// TIA Portal project "liquid refill system" (V18)

(* hardware
DEVICE "S7-1200 station_1"  S7-1200 Station
   slot 0: "Rack_0"  S7-1200 Rack  Rack  V1.0
   slot 1: "PLC_Refill"  CPU 1214C DC/DC/Rly  6ES7 214-1HG40-0XB0  V4.6
DEVICE "HMI_Refill"  TP900 Comfort
   slot 0: "HMI_Refill"  TP900 Comfort  6AV2 124-0JC01-0AX0  17.0.0.0
   slot 1: "HMI_RT_1"  TP900 Comfort  6AV2 124-0JC01-0AX0  17.0.0.0
   slot 5: "HMI_Refill.IE_CP_1"  PROFINET Interface  17.0.0.0
      slot 1: "PROFINET Interface_1"  PROFINET Interface
         slot 1: "Port_1"  Port
         slot 2: "Port_2"  Port
   slot 7: "HMI_Refill.MPI/DP_CP_1"  MPI/DP Interface  17.0.0.0
*)

// ===== PLC "PLC_Refill"  CPU 1214C DC/DC/Rly =====

VAR_GLOBAL   // PLC tag table "Default tag table"
   "System_Byte" AT %MB1 : Byte;
   "FirstScan" AT %M1.0 : Bool;
   "DiagStatusUpdate" AT %M1.1 : Bool;
   "AlwaysTRUE" AT %M1.2 : Bool;
   "AlwaysFALSE" AT %M1.3 : Bool;
   "Clock_Byte" AT %MB0 : Byte;
   "Clock_10Hz" AT %M0.0 : Bool;
   "Clock_5Hz" AT %M0.1 : Bool;
   "Clock_2.5Hz" AT %M0.2 : Bool;
   "Clock_2Hz" AT %M0.3 : Bool;
   "Clock_1.25Hz" AT %M0.4 : Bool;
   "Clock_1Hz" AT %M0.5 : Bool;
   "Clock_0.625Hz" AT %M0.6 : Bool;
   "Clock_0.5Hz" AT %M0.7 : Bool;
END_VAR

VAR_GLOBAL   // PLC tag table "input Machine"
   "i_Start" AT %I0.0 : Bool;
   "i_Stop" AT %I0.1 : Bool;
   "i_Reset" AT %I0.2 : Bool;
END_VAR

VAR_GLOBAL   // PLC tag table "output Machine"
   "q_Lamp_Running" AT %Q0.0 : Bool;   // Indication lamp, application running
   "q_Lamp_Faulted" AT %Q0.1 : Bool;   // Indication lamp, application faulted
   "q_Lamp_Ready" AT %Q0.7 : Bool;   // Indication lamp, application ready
END_VAR

VAR_GLOBAL   // PLC tag table "input Equipment"
   "iw_RefillTank1_Level" AT %IW64 : Int;   // Refill tank actual water level process
   "iw_RefillTank2_Level" AT %IW66 : Int;   // Refill tank actual water level process
   "i_RefillPump1_MCB" AT %I0.3 : Bool;   // Refill pump motor circuit breaker process ( Motor saftety )
   "i_RefillPump1_LI" AT %I0.4 : Bool;   // Refill pump local isolator process( Human safety )
   "i_RefillPump1_running" AT %I0.5 : Bool;   // Refill Pump Running feedback
   "i_RefillValve1_feedback" AT %I0.6 : Bool;   // Refill Valve position open feedback
   "i_RefillPump2_MCB" AT %I0.7 : Bool;   // Refill pump motor circuit breaker process ( Motor saftety )
   "i_RefillPump2_LI" AT %I1.0 : Bool;   // Refill pump local isolator process( Human safety )
   "i_RefillPump2_running" AT %I1.1 : Bool;   // Refill Pump Running feedback
   "i_RefillValve2_feedback" AT %I1.2 : Bool;   // Refill Valve position open feedback
   "i_SupplyTank_lowlevel" AT %I1.3 : Bool;   // Supply tank low level indicator
   "i_SupplyValve_feedback" AT %I1.4 : Bool;   // Supply valve position open feedback
END_VAR

VAR_GLOBAL   // PLC tag table "output Equipment"
   "q_RefillPump1_Start" AT %Q0.2 : Bool;   // Refill pump start operation process
   "q_RefillValve1_Open" AT %Q0.3 : Bool;   // Refill valve open operation process
   "q_RefillPump2_Start" AT %Q0.4 : Bool;   // Refill pump start operation process
   "q_RefillValve2_Open" AT %Q0.5 : Bool;   // Refill valve open operation process
   "q_SupplyValve_Open" AT %Q0.6 : Bool;   // Supply valve open operation process
END_VAR

TYPE "UDT_Statehandler"
   STRUCT
      State : Struct   // System states
         iState : Int;   // State feedback
         xReady : Bool;   // System is in ready state
         xRunning : Bool;   // System is in running state
         xFaulted : Bool;   // System is in faulted state
         xReset : Bool;   // System is in reset fault state
      END_STRUCT;
      Cmd : Struct   // Command structure
         xStart : Bool;   // Start operation - button on HMI
         xStop : Bool;   // Stop operation - button on HMI
         xReset : Bool;   // Reset faults - button on HMI
      END_STRUCT;
   END_STRUCT;
END_TYPE

TYPE "UDT_Refill"
   STRUCT
      Sts : Struct   // Status structure
         iTankLevel : Int;   // Actual product level in tank
         iPumpState : Int;   // Pump state (0=off,1=running,2=faulted)
         iValveState : Int;   // Valve state (0=closed,1=open,2=faulted)
         xPumpRunning : Bool;   // Pump is in operation
         xValveOpen : Bool;   // Valve is in open position
         xFaulted : Bool;   // Refill system faulted
      END_STRUCT;
      Cmd : Struct   // Command structure
         xRequestRefill : Bool;   // Request a refill
      END_STRUCT;
      Par : Struct   // Parameter structure
         iTankLevelLow : Int;   // Tank low level (%)
         iTankLevelHigh : Int;   // Tank high level (%)
      END_STRUCT;
      Cfg : Struct   // Configuration structure
         xSpare : Bool;   // spare ( reserve )
      END_STRUCT;
      Flt : Struct   // Fault Structure
         wTrigger : Word;   // Fault triggers
      END_STRUCT;
   END_STRUCT;
END_TYPE

TYPE "UDT_Supply"
   STRUCT
      Sts : Struct   // Status structure
         iValveState : Int;   // Valve state (0=closed,1=open,2=faulted)
         xTankLowLevel : Bool;   // Low product level in tank
         xValveOpen : Bool;   // Valve is in open position
         xFaulted : Bool;   // Supply system faulted
      END_STRUCT;
      Cmd : Struct   // Command structure
         xSpare : Bool;   // spare(reserve)
      END_STRUCT;
      Par : Struct   // Parameter structure
         rTankLowLevelDelay : Real;   // rTankLowLevelDelay
      END_STRUCT;
      Cfg : Struct   // Configuration structure
         xSpare : Bool;   // spare(reserve)
      END_STRUCT;
      Flt : Struct   // Fault structure
         wTrigger : Word;   // Fault triggers
      END_STRUCT;
   END_STRUCT;
END_TYPE

// folder: 00 Machine

DATA_BLOCK "Instance_Machine Module"   // DB4
{ S7_Optimized_Access := 'TRUE' }
VERSION : 0.1
// stored: InstanceOfName FB_Machine Module
"FB_Machine Module"
BEGIN
END_DATA_BLOCK

// folder: 01 Equipment

DATA_BLOCK "FB_Equipment Modules_DB"   // DB5
{ S7_Optimized_Access := 'TRUE' }
VERSION : 0.1
// stored: InstanceOfName FB_Equipment Modules
"FB_Equipment Modules"
BEGIN
END_DATA_BLOCK

// folder: Global DB

DATA_BLOCK "DB - Machine"   // DB1
{ S7_Optimized_Access := 'TRUE' }
VERSION : 0.1
   VAR
      StateHandler : "UDT_Statehandler";
   END_VAR
BEGIN
END_DATA_BLOCK

DATA_BLOCK "DB - Equipment"   // DB2
{ S7_Optimized_Access := 'TRUE' }
VERSION : 0.1
   VAR
      Supply : "UDT_Supply";
      Refill_Process_1 : "UDT_Refill";
      Refill_Process_2 : "UDT_Refill";
   END_VAR
BEGIN
END_DATA_BLOCK

// folder: (top level)

ORGANIZATION_BLOCK "Main"   // OB1, LAD, ProgramCycle
TITLE = "Main Program Sweep (Cycle)"
{ S7_Optimized_Access := 'TRUE' }
VERSION : 0.1
   VAR_INPUT
      Initial_Call : Bool;   // Initial call of this OB
      Remanence : Bool;   // =True, if remanent data are available
   END_VAR
BEGIN

REGION Network 1: CALL - Main machine modules
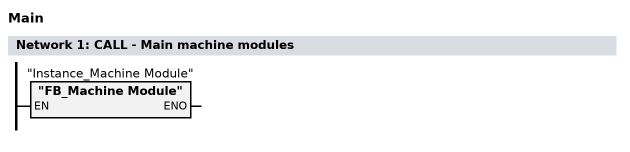
   RUNG wire#powerrail
      "Instance_Machine Module"()
   END_RUNG
   // the same network as SCL:
   "Instance_Machine Module"();   // "FB_Machine Module"
END_REGION

REGION Network 2: CALL - Main equipment modules
END_REGION
END_ORGANIZATION_BLOCK

// folder: 00 Machine

FUNCTION_BLOCK "FB_Machine Module"   // FB1, LAD
{ S7_Optimized_Access := 'TRUE' }
VERSION : 0.1
   VAR
      FB_StateHandler_Instance : "FB_StateHandler";
   END_VAR
   VAR_TEMP
      info : Struct
         xReady : Bool;
         xRunning : Bool;
         xFaulted : Bool;
         xReset : Bool;
      END_STRUCT;
   END_VAR
BEGIN

REGION Network 1
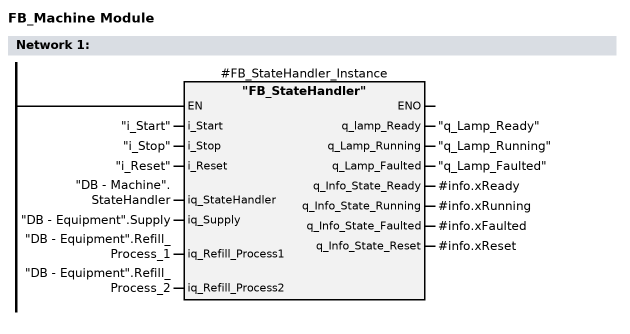
   RUNG wire#powerrail
      #FB_StateHandler_Instance(i_Start := "i_Start", i_Stop := "i_Stop", i_Reset := "i_Reset", iq_StateHandler := "DB - Machine".StateHandler, iq_Supply := "DB - Equipment".Supply, iq_Refill_Process1 := "DB - Equipment".Refill_Process_1, iq_Refill_Process2 := "DB - Equipment".Refill_Process_2, q_lamp_Ready => "q_Lamp_Ready", q_Lamp_Running => "q_Lamp_Running", q_Lamp_Faulted => "q_Lamp_Faulted", q_Info_State_Ready => #info.xReady, q_Info_State_Running => #info.xRunning, q_Info_State_Faulted => #info.xFaulted, q_Info_State_Reset => #info.xReset)
   END_RUNG
   // the same network as SCL:
   #FB_StateHandler_Instance(i_Start := "i_Start",   // "FB_StateHandler"
                           i_Stop := "i_Stop",
                           i_Reset := "i_Reset",
                           iq_StateHandler := "DB - Machine".StateHandler,
                           iq_Supply := "DB - Equipment".Supply,
                           iq_Refill_Process1 := "DB - Equipment".Refill_Process_1,
                           iq_Refill_Process2 := "DB - Equipment".Refill_Process_2,
                           q_lamp_Ready => "q_Lamp_Ready",
                           q_Lamp_Running => "q_Lamp_Running",
                           q_Lamp_Faulted => "q_Lamp_Faulted",
                           q_Info_State_Ready => #info.xReady,
                           q_Info_State_Running => #info.xRunning,
                           q_Info_State_Faulted => #info.xFaulted,
                           q_Info_State_Reset => #info.xReset);
END_REGION
END_FUNCTION_BLOCK

// folder: 00 Machine/Function

FUNCTION_BLOCK "FB_StateHandler"   // FB2, LAD
TITLE = MACHINE - State Handler
{ S7_Optimized_Access := 'TRUE' }
VERSION : 0.1
// This function block contains all logic for control and status of the machine state handler.
// This module consists of 4 states: start, stop, faulted and reset.
   VAR_INPUT
      i_Start : Bool;
      i_Stop : Bool;
      i_Reset : Bool;
   END_VAR
   VAR_OUTPUT
      q_lamp_Ready : Bool;
      q_Lamp_Running : Bool;   // Lamp machine running
      q_Lamp_Faulted : Bool;   // Lamp machine faulted
      q_Info_State_Ready : Bool;
      q_Info_State_Running : Bool;
      q_Info_State_Faulted : Bool;
      q_Info_State_Reset : Bool;
   END_VAR
   VAR_IN_OUT
      iq_StateHandler : "UDT_Statehandler";
      iq_Supply : "UDT_Supply";
      iq_Refill_Process1 : "UDT_Refill";
      iq_Refill_Process2 : "UDT_Refill";
   END_VAR
   VAR
      stOnDelay_Reset : IEC_TIMER;
      iState : Int;
   END_VAR
   VAR_TEMP
      _tTimeET : Time;
   END_VAR
BEGIN

REGION Network 1: CONTROL - Start Operation
   // The application goes from a ready state (0) to a running state (1) by pressing Start
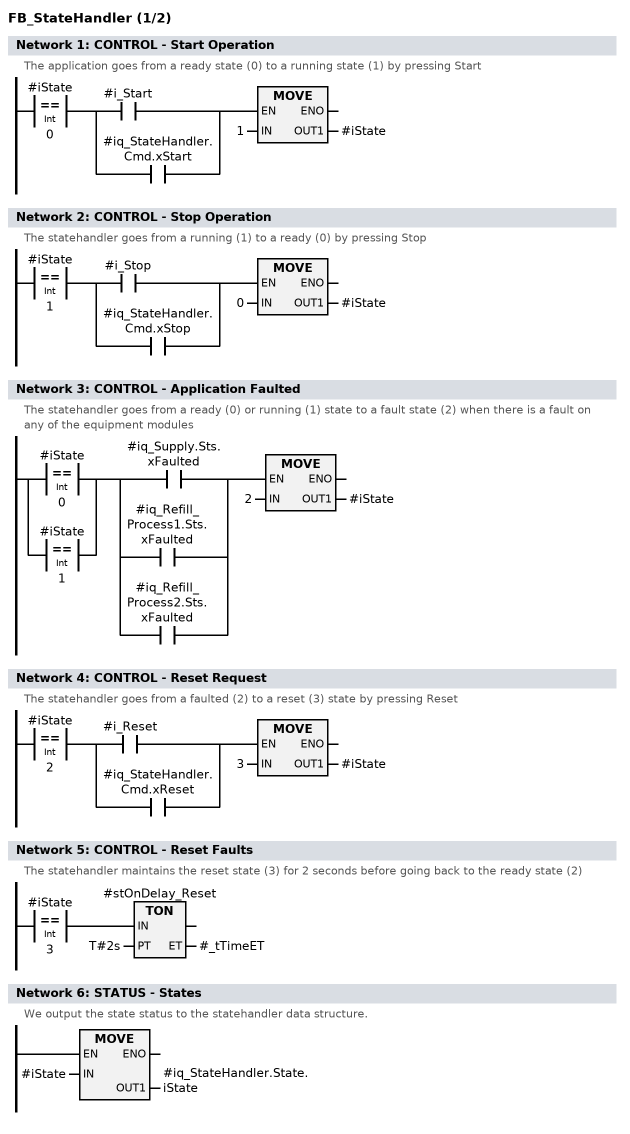
   RUNG wire#powerrail
      { S7_Templates := "SrcType := Int" } EQ_Contact(in1 := #iState, in2 := 0)
      wire#w1
      Contact( #i_Start )
      wire#w2
      Move(in := 1, out1 => #iState)
   END_RUNG
   RUNG wire#w1
      Contact( #iq_StateHandler.Cmd.xStart )
   END_RUNG wire#w2
   // the same network as SCL:
   IF (#iState = 0) AND (#i_Start OR #iq_StateHandler.Cmd.xStart) THEN #iState := 1; END_IF;
END_REGION

REGION Network 2: CONTROL - Stop Operation
   // The statehandler goes from a running (1) to a ready (0) by pressing Stop
   RUNG wire#powerrail
      { S7_Templates := "SrcType := Int" } EQ_Contact(in1 := #iState, in2 := 1)
      wire#w1
      Contact( #i_Stop )
      wire#w2
      Move(in := 0, out1 => #iState)
   END_RUNG
   RUNG wire#w1
      Contact( #iq_StateHandler.Cmd.xStop )
   END_RUNG wire#w2
   // the same network as SCL:
   IF (#iState = 1) AND (#i_Stop OR #iq_StateHandler.Cmd.xStop) THEN #iState := 0; END_IF;
END_REGION

REGION Network 3: CONTROL - Application Faulted
   // The statehandler goes from a ready (0) or running (1) state to a fault state (2) when there is a fault on any of the equipment modules
   RUNG wire#powerrail
      { S7_Templates := "SrcType := Int" } EQ_Contact(in1 := #iState, in2 := 0)
      wire#w1
      Contact( #iq_Supply.Sts.xFaulted )
      wire#w2
      Move(in := 2, out1 => #iState)
   END_RUNG
   RUNG wire#powerrail
      { S7_Templates := "SrcType := Int" } EQ_Contact(in1 := #iState, in2 := 1)
   END_RUNG wire#w1
   RUNG wire#w1
      Contact( #iq_Refill_Process1.Sts.xFaulted )
   END_RUNG wire#w2
   RUNG wire#w1
      Contact( #iq_Refill_Process2.Sts.xFaulted )
   END_RUNG wire#w2
   // the same network as SCL:
   IF ((#iState = 0) OR (#iState = 1)) AND (#iq_Supply.Sts.xFaulted OR #iq_Refill_Process1.Sts.xFaulted OR #iq_Refill_Process2.Sts.xFaulted) THEN
       #iState := 2;
   END_IF;
END_REGION

REGION Network 4: CONTROL - Reset Request
   // The statehandler goes from a faulted (2) to a reset (3) state by pressing Reset
   RUNG wire#powerrail
      { S7_Templates := "SrcType := Int" } EQ_Contact(in1 := #iState, in2 := 2)
      wire#w1
      Contact( #i_Reset )
      wire#w2
      Move(in := 3, out1 => #iState)
   END_RUNG
   RUNG wire#w1
      Contact( #iq_StateHandler.Cmd.xReset )
   END_RUNG wire#w2
   // the same network as SCL:
   IF (#iState = 2) AND (#i_Reset OR #iq_StateHandler.Cmd.xReset) THEN #iState := 3; END_IF;
END_REGION

REGION Network 5: CONTROL - Reset Faults
   // The statehandler maintains the reset state (3) for 2 seconds before going back to the ready state (2)
   #stOnDelay_Reset.TON(IN := #iState = 3, PT := T#2s, ET => #_tTimeET);
END_REGION

REGION Network 6: STATUS - States
   // We output the state status to the statehandler data structure.
   RUNG wire#powerrail
      Move(in := #iState, out1 => #iq_StateHandler.State.iState)
   END_RUNG
   // the same network as SCL:
   #iq_StateHandler.State.iState := #iState;
END_REGION

REGION Network 7: STATUS - State Ready
   // The ready state is defined by state "0". We output the ready state status to the statehandler data structure and as an information output on the block.
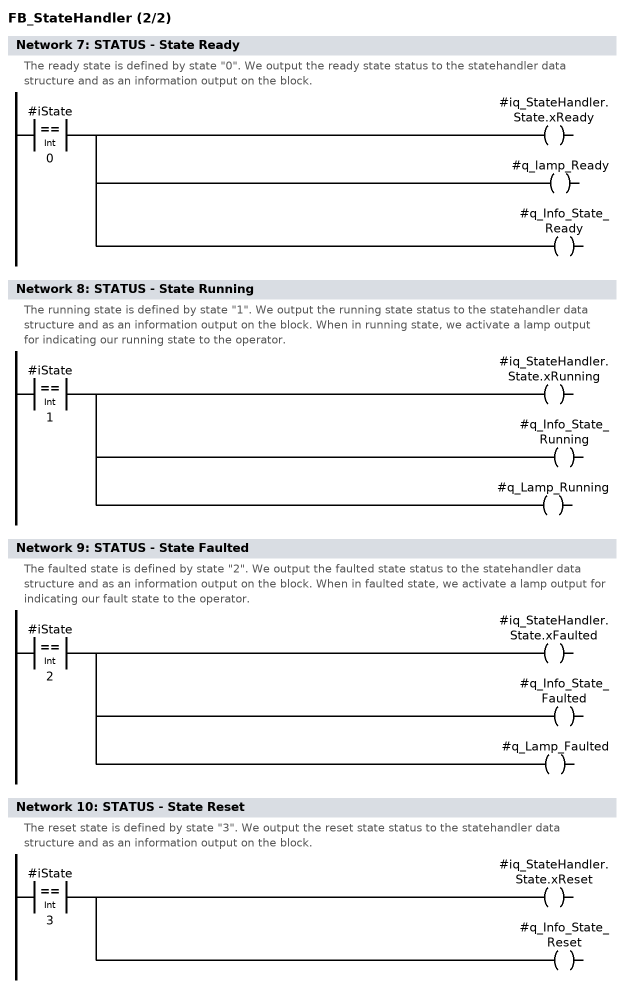
   RUNG wire#powerrail
      { S7_Templates := "SrcType := Int" } EQ_Contact(in1 := #iState, in2 := 0)
      wire#w1
      Coil( #iq_StateHandler.State.xReady )
   END_RUNG
   RUNG wire#w1
      Coil( #q_lamp_Ready )
   END_RUNG
   RUNG wire#w1
      Coil( #q_Info_State_Ready )
   END_RUNG
   // the same network as SCL:
   #iq_StateHandler.State.xReady := #iState = 0;
   #q_lamp_Ready := #iq_StateHandler.State.xReady;
   #q_Info_State_Ready := #iq_StateHandler.State.xReady;
END_REGION

REGION Network 8: STATUS - State Running
   // The running state is defined by state "1". We output the running state status to the statehandler data structure and as an information output on the block. When in running state, we activate a lamp output for indicating our running state to the operator.
   RUNG wire#powerrail
      { S7_Templates := "SrcType := Int" } EQ_Contact(in1 := #iState, in2 := 1)
      wire#w1
      Coil( #iq_StateHandler.State.xRunning )
   END_RUNG
   RUNG wire#w1
      Coil( #q_Info_State_Running )
   END_RUNG
   RUNG wire#w1
      Coil( #q_Lamp_Running )
   END_RUNG
   // the same network as SCL:
   #iq_StateHandler.State.xRunning := #iState = 1;
   #q_Info_State_Running := #iq_StateHandler.State.xRunning;
   #q_Lamp_Running := #iq_StateHandler.State.xRunning;
END_REGION

REGION Network 9: STATUS - State Faulted
   // The faulted state is defined by state "2". We output the faulted state status to the statehandler data structure and as an information output on the block. When in faulted state, we activate a lamp output for indicating our fault state to the operator.
   RUNG wire#powerrail
      { S7_Templates := "SrcType := Int" } EQ_Contact(in1 := #iState, in2 := 2)
      wire#w1
      Coil( #iq_StateHandler.State.xFaulted )
   END_RUNG
   RUNG wire#w1
      Coil( #q_Info_State_Faulted )
   END_RUNG
   RUNG wire#w1
      Coil( #q_Lamp_Faulted )
   END_RUNG
   // the same network as SCL:
   #iq_StateHandler.State.xFaulted := #iState = 2;
   #q_Info_State_Faulted := #iq_StateHandler.State.xFaulted;
   #q_Lamp_Faulted := #iq_StateHandler.State.xFaulted;
END_REGION

REGION Network 10: STATUS - State Reset
   // The reset state is defined by state "3". We output the reset state status to the statehandler data structure and as an information output on the block.
   RUNG wire#powerrail
      { S7_Templates := "SrcType := Int" } EQ_Contact(in1 := #iState, in2 := 3)
      wire#w1
      Coil( #iq_StateHandler.State.xReset )
   END_RUNG
   RUNG wire#w1
      Coil( #q_Info_State_Reset )
   END_RUNG
   // the same network as SCL:
   #iq_StateHandler.State.xReset := #iState = 3;
   #q_Info_State_Reset := #iq_StateHandler.State.xReset;
END_REGION
END_FUNCTION_BLOCK

// folder: 01 Equipment

FUNCTION_BLOCK "FB_Equipment Modules"   // FB3, LAD
{ S7_Optimized_Access := 'TRUE' }
VERSION : 0.1
   VAR
      FB_Supply_Instance : "FB_Supply";
      FB_Refill_Instance : "FB_Refill";
      FB_Refill_Instance_1 : "FB_Refill";
   END_VAR
   VAR_TEMP
      Info_FaultedSupply : Bool;
      info_FaultedRefill1 : Bool;
      info_FaultedRefill2 : Bool;
   END_VAR
BEGIN

REGION Network 1: MODULE - Supply
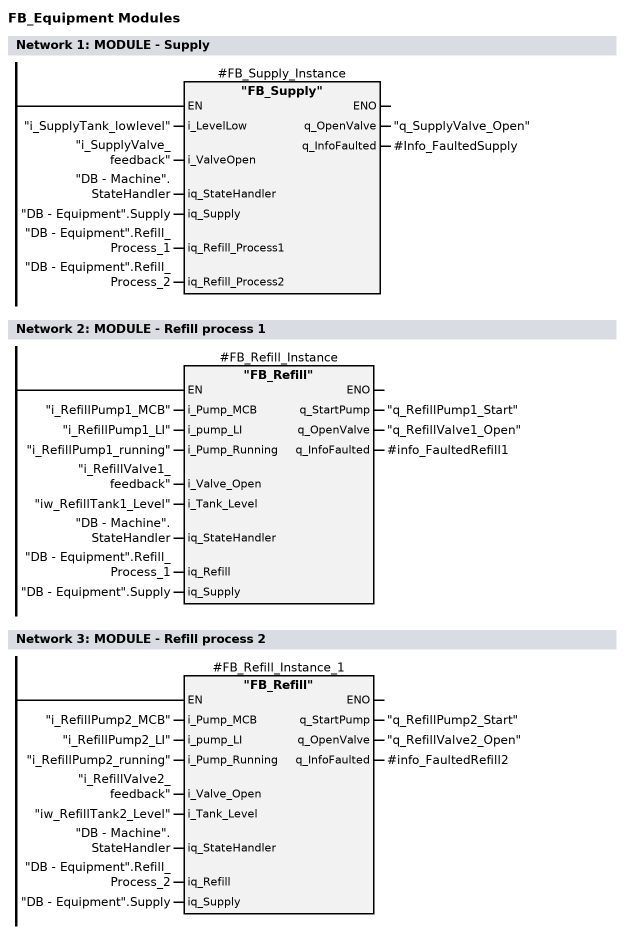
   RUNG wire#powerrail
      #FB_Supply_Instance(i_LevelLow := "i_SupplyTank_lowlevel", i_ValveOpen := "i_SupplyValve_feedback", iq_StateHandler := "DB - Machine".StateHandler, iq_Supply := "DB - Equipment".Supply, iq_Refill_Process1 := "DB - Equipment".Refill_Process_1, iq_Refill_Process2 := "DB - Equipment".Refill_Process_2, q_OpenValve => "q_SupplyValve_Open", q_InfoFaulted => #Info_FaultedSupply)
   END_RUNG
   // the same network as SCL:
   #FB_Supply_Instance(i_LevelLow := "i_SupplyTank_lowlevel",   // "FB_Supply"
                       i_ValveOpen := "i_SupplyValve_feedback",
                       iq_StateHandler := "DB - Machine".StateHandler,
                       iq_Supply := "DB - Equipment".Supply,
                       iq_Refill_Process1 := "DB - Equipment".Refill_Process_1,
                       iq_Refill_Process2 := "DB - Equipment".Refill_Process_2,
                       q_OpenValve => "q_SupplyValve_Open",
                       q_InfoFaulted => #Info_FaultedSupply);
END_REGION

REGION Network 2: MODULE - Refill process 1
   RUNG wire#powerrail
      #FB_Refill_Instance(i_Pump_MCB := "i_RefillPump1_MCB", i_pump_LI := "i_RefillPump1_LI", i_Pump_Running := "i_RefillPump1_running", i_Valve_Open := "i_RefillValve1_feedback", i_Tank_Level := "iw_RefillTank1_Level", iq_StateHandler := "DB - Machine".StateHandler, iq_Refill := "DB - Equipment".Refill_Process_1, iq_Supply := "DB - Equipment".Supply, q_StartPump => "q_RefillPump1_Start", q_OpenValve => "q_RefillValve1_Open", q_InfoFaulted => #info_FaultedRefill1)
   END_RUNG
   // the same network as SCL:
   #FB_Refill_Instance(i_Pump_MCB := "i_RefillPump1_MCB",   // "FB_Refill"
                       i_pump_LI := "i_RefillPump1_LI",
                       i_Pump_Running := "i_RefillPump1_running",
                       i_Valve_Open := "i_RefillValve1_feedback",
                       i_Tank_Level := "iw_RefillTank1_Level",
                       iq_StateHandler := "DB - Machine".StateHandler,
                       iq_Refill := "DB - Equipment".Refill_Process_1,
                       iq_Supply := "DB - Equipment".Supply,
                       q_StartPump => "q_RefillPump1_Start",
                       q_OpenValve => "q_RefillValve1_Open",
                       q_InfoFaulted => #info_FaultedRefill1);
END_REGION

REGION Network 3: MODULE - Refill process 2
   RUNG wire#powerrail
      #FB_Refill_Instance_1(i_Pump_MCB := "i_RefillPump2_MCB", i_pump_LI := "i_RefillPump2_LI", i_Pump_Running := "i_RefillPump2_running", i_Valve_Open := "i_RefillValve2_feedback", i_Tank_Level := "iw_RefillTank2_Level", iq_StateHandler := "DB - Machine".StateHandler, iq_Refill := "DB - Equipment".Refill_Process_2, iq_Supply := "DB - Equipment".Supply, q_StartPump => "q_RefillPump2_Start", q_OpenValve => "q_RefillValve2_Open", q_InfoFaulted => #info_FaultedRefill2)
   END_RUNG
   // the same network as SCL:
   #FB_Refill_Instance_1(i_Pump_MCB := "i_RefillPump2_MCB",   // "FB_Refill"
                         i_pump_LI := "i_RefillPump2_LI",
                         i_Pump_Running := "i_RefillPump2_running",
                         i_Valve_Open := "i_RefillValve2_feedback",
                         i_Tank_Level := "iw_RefillTank2_Level",
                         iq_StateHandler := "DB - Machine".StateHandler,
                         iq_Refill := "DB - Equipment".Refill_Process_2,
                         iq_Supply := "DB - Equipment".Supply,
                         q_StartPump => "q_RefillPump2_Start",
                         q_OpenValve => "q_RefillValve2_Open",
                         q_InfoFaulted => #info_FaultedRefill2);
END_REGION
END_FUNCTION_BLOCK

// folder: 01 Equipment/Function

FUNCTION_BLOCK "FB_Refill"   // FB4, LAD
TITLE = EQUIPMENT - Refill
{ S7_Optimized_Access := 'TRUE' }
VERSION : 0.1
// This module consists of a tank with an analog level sensor, a pump and a valve.
   VAR_INPUT
      i_Pump_MCB : Bool;
      i_pump_LI : Bool;
      i_Pump_Running : Bool;
      i_Valve_Open : Bool;
      i_Tank_Level : Int;
   END_VAR
   VAR_OUTPUT
      q_StartPump : Bool;
      q_OpenValve : Bool;
      q_InfoFaulted : Bool;
   END_VAR
   VAR_IN_OUT
      iq_StateHandler : "UDT_Statehandler";
      iq_Refill : "UDT_Refill";
      iq_Supply : "UDT_Supply";
   END_VAR
   VAR
      OnDelay_Flt_Pump_Running : IEC_TIMER;
      OnDelay_Flt_Valve_Open : IEC_TIMER;
   END_VAR
   VAR_TEMP
      Cmd_StartPump : Bool;
      Cmd_OpenValve : Bool;
      TimeET : Time;
      Flt_Pump : Bool;
      Flt_Valve : Bool;
   END_VAR
BEGIN

REGION Network 1: REQUEST - Refill
   // Start refilling when tank level goes below 10%.
   // Stop refilling when tank level goes above 60%.
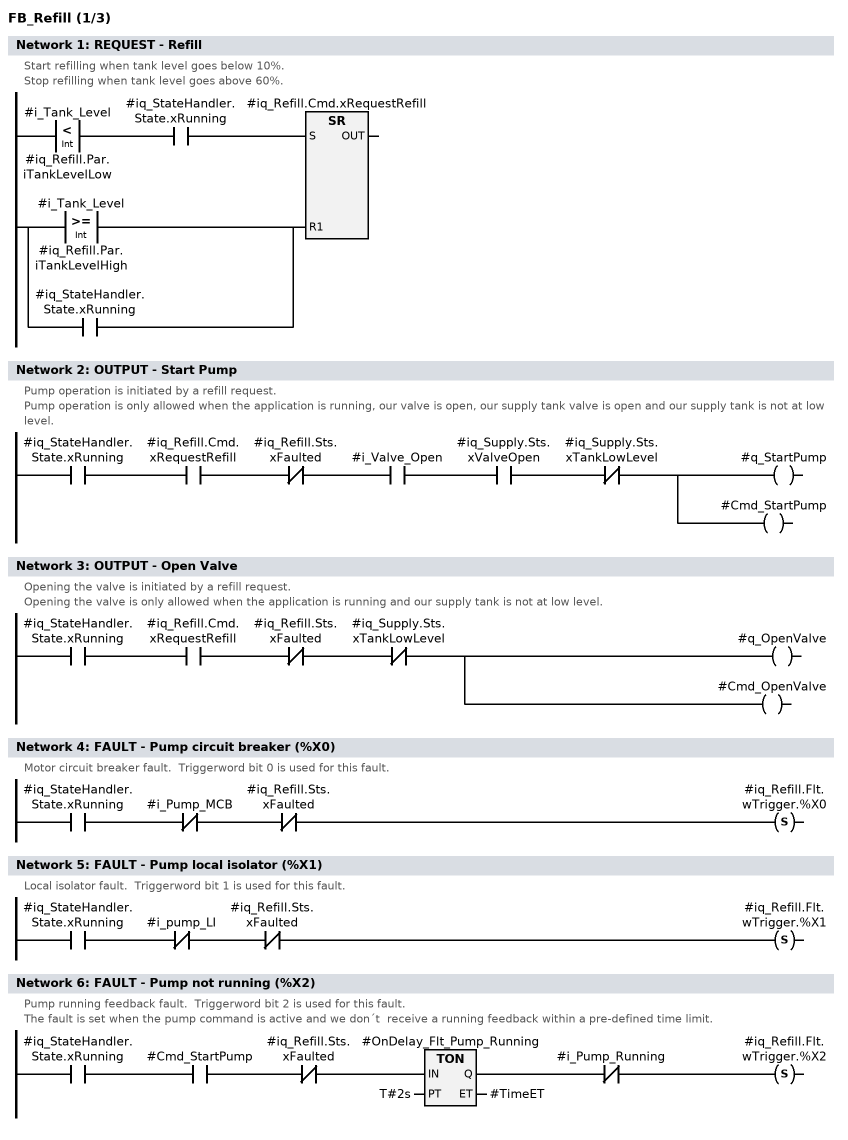
   RUNG wire#powerrail
      { S7_Templates := "SrcType := Int" } LT_Contact(in1 := #i_Tank_Level, in2 := #iq_Refill.Par.iTankLevelLow)
      Contact( #iq_StateHandler.State.xRunning )
      S_SR(operand := #iq_Refill.Cmd.xRequestRefill, r1 := wire#w1)
   END_RUNG
   RUNG wire#powerrail
      { S7_Templates := "SrcType := Int" } GE_Contact(in1 := #i_Tank_Level, in2 := #iq_Refill.Par.iTankLevelHigh)
   END_RUNG wire#w1
   RUNG wire#powerrail
      Contact( #iq_StateHandler.State.xRunning )
   END_RUNG wire#w1
   // the same network as SCL:
   IF (#i_Tank_Level < #iq_Refill.Par.iTankLevelLow) AND #iq_StateHandler.State.xRunning THEN
       #iq_Refill.Cmd.xRequestRefill := TRUE;   // SR flip-flop
   END_IF;
   IF (#i_Tank_Level >= #iq_Refill.Par.iTankLevelHigh) OR #iq_StateHandler.State.xRunning THEN
       #iq_Refill.Cmd.xRequestRefill := FALSE;
   END_IF;
END_REGION

REGION Network 2: OUTPUT - Start Pump
   // Pump operation is initiated by a refill request.
   // Pump operation is only allowed when the application is running, our valve is open, our supply tank valve is open and our supply tank is not at low level.
   RUNG wire#powerrail
      Contact( #iq_StateHandler.State.xRunning )
      Contact( #iq_Refill.Cmd.xRequestRefill )
      I_Contact( #iq_Refill.Sts.xFaulted )
      Contact( #i_Valve_Open )
      Contact( #iq_Supply.Sts.xValveOpen )
      I_Contact( #iq_Supply.Sts.xTankLowLevel )
      wire#w1
      Coil( #q_StartPump )
   END_RUNG
   RUNG wire#w1
      Coil( #Cmd_StartPump )
   END_RUNG
   // the same network as SCL:
   #q_StartPump := #iq_StateHandler.State.xRunning AND #iq_Refill.Cmd.xRequestRefill AND NOT #iq_Refill.Sts.xFaulted AND #i_Valve_Open AND #iq_Supply.Sts.xValveOpen AND NOT #iq_Supply.Sts.xTankLowLevel;
   #Cmd_StartPump := #q_StartPump;
END_REGION

REGION Network 3: OUTPUT - Open Valve
   // Opening the valve is initiated by a refill request.
   // Opening the valve is only allowed when the application is running and our supply tank is not at low level.
   RUNG wire#powerrail
      Contact( #iq_StateHandler.State.xRunning )
      Contact( #iq_Refill.Cmd.xRequestRefill )
      I_Contact( #iq_Refill.Sts.xFaulted )
      I_Contact( #iq_Supply.Sts.xTankLowLevel )
      wire#w1
      Coil( #q_OpenValve )
   END_RUNG
   RUNG wire#w1
      Coil( #Cmd_OpenValve )
   END_RUNG
   // the same network as SCL:
   #q_OpenValve := #iq_StateHandler.State.xRunning AND #iq_Refill.Cmd.xRequestRefill AND NOT #iq_Refill.Sts.xFaulted AND NOT #iq_Supply.Sts.xTankLowLevel;
   #Cmd_OpenValve := #q_OpenValve;
END_REGION

REGION Network 4: FAULT - Pump circuit breaker (%X0)
   // Motor circuit breaker fault.  Triggerword bit 0 is used for this fault.
   RUNG wire#powerrail
      Contact( #iq_StateHandler.State.xRunning )
      I_Contact( #i_Pump_MCB )
      I_Contact( #iq_Refill.Sts.xFaulted )
      S_Coil( #iq_Refill.Flt.wTrigger.%X0 )
   END_RUNG
   // the same network as SCL:
   IF #iq_StateHandler.State.xRunning AND NOT #i_Pump_MCB AND NOT #iq_Refill.Sts.xFaulted THEN
       #iq_Refill.Flt.wTrigger.%X0 := TRUE;
   END_IF;
END_REGION

REGION Network 5: FAULT - Pump local isolator (%X1)
   // Local isolator fault.  Triggerword bit 1 is used for this fault.
   RUNG wire#powerrail
      Contact( #iq_StateHandler.State.xRunning )
      I_Contact( #i_pump_LI )
      I_Contact( #iq_Refill.Sts.xFaulted )
      S_Coil( #iq_Refill.Flt.wTrigger.%X1 )
   END_RUNG
   // the same network as SCL:
   IF #iq_StateHandler.State.xRunning AND NOT #i_pump_LI AND NOT #iq_Refill.Sts.xFaulted THEN
       #iq_Refill.Flt.wTrigger.%X1 := TRUE;
   END_IF;
END_REGION

REGION Network 6: FAULT - Pump not running (%X2)
   // Pump running feedback fault.  Triggerword bit 2 is used for this fault.
   // The fault is set when the pump command is active and we don´t  receive a running feedback within a pre-defined time limit.
   #OnDelay_Flt_Pump_Running.TON(IN := #iq_StateHandler.State.xRunning AND #Cmd_StartPump AND NOT #iq_Refill.Sts.xFaulted,
                           PT := T#2s,
                           ET => #TimeET);
   IF #OnDelay_Flt_Pump_Running.Q AND NOT #i_Pump_Running THEN #iq_Refill.Flt.wTrigger.%X2 := TRUE; END_IF;
END_REGION

REGION Network 7: FAULT - Valve not opening (%X3)
   // Valve open position fault.  Triggerword bit 3 is used for this fault.
   // The fault is set when the valve open command is active and we don´t  receive an open position feedback within a pre-defined time limit.